   "TT426STR_ALM_ANALOG_DB_VERY LOW LEVEL VALUE (LL)" : Real = PLC TT426STR_ALM_ANALOG_DB."VERY LOW LEVEL VALUE (LL)" AT %DB2072.DBD22, 1 s
   "IDB_TIT 360_VERY HIGH LEVEL VALUE (HH)" : Real = PLC "IDB_TIT 360"."VERY HIGH LEVEL VALUE (HH)" AT %DB760.DBD34, 1 s
   "IDB_TIT 360_HIGH LEVEL VALUE (H)" : Real = PLC "IDB_TIT 360"."HIGH LEVEL VALUE (H)" AT %DB760.DBD30, 1 s
   "IDB_TIT 360_LOW LEVEL VALUE (L)" : Real = PLC "IDB_TIT 360"."LOW LEVEL VALUE (L)" AT %DB760.DBD26, 1 s
   "IDB_TIT 360_VERY LOW LEVEL VALUE (LL)" : Real = PLC "IDB_TIT 360"."VERY LOW LEVEL VALUE (LL)" AT %DB760.DBD22, 1 s
   "IDB_TIT 319_VERY HIGH LEVEL VALUE (HH)" : Real = PLC "IDB_TIT 319"."VERY HIGH LEVEL VALUE (HH)" AT %DB719.DBD34, 1 s
   "IDB_TIT 319_HIGH LEVEL VALUE (H)" : Real = PLC "IDB_TIT 319"."HIGH LEVEL VALUE (H)" AT %DB719.DBD30, 1 s
   "IDB_TIT 319_LOW LEVEL VALUE (L)" : Real = PLC "IDB_TIT 319"."LOW LEVEL VALUE (L)" AT %DB719.DBD26, 1 s
   "IDB_TIT 319_VERY LOW LEVEL VALUE (LL)" : Real = PLC "IDB_TIT 319"."VERY LOW LEVEL VALUE (LL)" AT %DB719.DBD22, 1 s
   "IDB_PIT 316_VERY HIGH LEVEL VALUE (HH)" : Real = PLC "IDB_PIT 316"."VERY HIGH LEVEL VALUE (HH)" AT %DB716.DBD34, 1 s
   "IDB_PIT 316_HIGH LEVEL VALUE (H)" : Real = PLC "IDB_PIT 316"."HIGH LEVEL VALUE (H)" AT %DB716.DBD30, 1 s
   "IDB_PIT 316_LOW LEVEL VALUE (L)" : Real = PLC "IDB_PIT 316"."LOW LEVEL VALUE (L)" AT %DB716.DBD26, 1 s
   "IDB_PIT 316_VERY LOW LEVEL VALUE (LL)" : Real = PLC "IDB_PIT 316"."VERY LOW LEVEL VALUE (LL)" AT %DB716.DBD22, 1 s
   "IDB_PIT 359_VERY HIGH LEVEL VALUE (HH)" : Real = PLC "IDB_PIT 359"."VERY HIGH LEVEL VALUE (HH)" AT %DB759.DBD34, 1 s
   "IDB_PIT 359_HIGH LEVEL VALUE (H)" : Real = PLC "IDB_PIT 359"."HIGH LEVEL VALUE (H)" AT %DB759.DBD30, 1 s
   "IDB_PIT 359_LOW LEVEL VALUE (L)" : Real = PLC "IDB_PIT 359"."LOW LEVEL VALUE (L)" AT %DB759.DBD26, 1 s
   "IDB_PIT 359_VERY LOW LEVEL VALUE (LL)" : Real = PLC "IDB_PIT 359"."VERY LOW LEVEL VALUE (LL)" AT %DB759.DBD22, 1 s
   "IDB_ATO2B_1_VERY HIGH LEVEL VALUE (HH)" : Real = PLC IDB_ATO2B_1."VERY HIGH LEVEL VALUE (HH)" AT %DB731.DBD34, 1 s
   "IDB_ATO2B_1_HIGH LEVEL VALUE (H)" : Real = PLC IDB_ATO2B_1."HIGH LEVEL VALUE (H)" AT %DB731.DBD30, 1 s
   "IDB_ATO2B_1_LOW LEVEL VALUE (L)" : Real = PLC IDB_ATO2B_1."LOW LEVEL VALUE (L)" AT %DB731.DBD26, 1 s
   "IDB_ATO2B_1_VERY LOW LEVEL VALUE (LL)" : Real = PLC IDB_ATO2B_1."VERY LOW LEVEL VALUE (LL)" AT %DB731.DBD22, 1 s
   "TT426_5S_ALM_ANALOG_DB_VERY HIGH LEVEL VALUE (HH)" : Real = PLC TT426_5S_ALM_ANALOG_DB."VERY HIGH LEVEL VALUE (HH)" AT %DB2082.DBD34, 1 s
   "TT426_5S_ALM_ANALOG_DB_HIGH LEVEL VALUE (H)" : Real = PLC TT426_5S_ALM_ANALOG_DB."HIGH LEVEL VALUE (H)" AT %DB2082.DBD30, 1 s
   "TT426_5S_ALM_ANALOG_DB_LOW LEVEL VALUE (L)" : Real = PLC TT426_5S_ALM_ANALOG_DB."LOW LEVEL VALUE (L)" AT %DB2082.DBD26, 1 s
   "TT426_5S_ALM_ANALOG_DB_VERY LOW LEVEL VALUE (LL)" : Real = PLC TT426_5S_ALM_ANALOG_DB."VERY LOW LEVEL VALUE (LL)" AT %DB2082.DBD22, 1 s
   "PIT424_RIO6_ALM_ANALOG_DB_VERY HIGH LEVEL VALUE (HH)" : Real = PLC PIT424_RIO6_ALM_ANALOG_DB."VERY HIGH LEVEL VALUE (HH)" AT %DB2223.DBD34, 1 s
   "PIT424_RIO6_ALM_ANALOG_DB_HIGH LEVEL VALUE (H)" : Real = PLC PIT424_RIO6_ALM_ANALOG_DB."HIGH LEVEL VALUE (H)" AT %DB2223.DBD30, 1 s
   "PIT424_RIO6_ALM_ANALOG_DB_LOW LEVEL VALUE (L)" : Real = PLC PIT424_RIO6_ALM_ANALOG_DB."LOW LEVEL VALUE (L)" AT %DB2223.DBD26, 1 s
   "PIT424_RIO6_ALM_ANALOG_DB_VERY LOW LEVEL VALUE (LL)" : Real = PLC PIT424_RIO6_ALM_ANALOG_DB."VERY LOW LEVEL VALUE (LL)" AT %DB2223.DBD22, 1 s
   "TT426_6P_ALM_ANALOG_DB_VERY HIGH LEVEL VALUE (HH)" : Real = PLC TT426_6P_ALM_ANALOG_DB."VERY HIGH LEVEL VALUE (HH)" AT %DB2083.DBD34, 1 s
   "TT426_6P_ALM_ANALOG_DB_HIGH LEVEL VALUE (H)" : Real = PLC TT426_6P_ALM_ANALOG_DB."HIGH LEVEL VALUE (H)" AT %DB2083.DBD30, 1 s
   "TT426_6P_ALM_ANALOG_DB_LOW LEVEL VALUE (L)" : Real = PLC TT426_6P_ALM_ANALOG_DB."LOW LEVEL VALUE (L)" AT %DB2083.DBD26, 1 s
   "TT426_6P_ALM_ANALOG_DB_VERY LOW LEVEL VALUE (LL)" : Real = PLC TT426_6P_ALM_ANALOG_DB."VERY LOW LEVEL VALUE (LL)" AT %DB2083.DBD22, 1 s
   "TT426_6S_ALM_ANALOG_DB_VERY HIGH LEVEL VALUE (HH)" : Real = PLC TT426_6S_ALM_ANALOG_DB."VERY HIGH LEVEL VALUE (HH)" AT %DB2085.DBD34, 1 s
   "TT426_6S_ALM_ANALOG_DB_HIGH LEVEL VALUE (H)" : Real = PLC TT426_6S_ALM_ANALOG_DB."HIGH LEVEL VALUE (H)" AT %DB2085.DBD30, 1 s
   "TT426_6S_ALM_ANALOG_DB_LOW LEVEL VALUE (L)" : Real = PLC TT426_6S_ALM_ANALOG_DB."LOW LEVEL VALUE (L)" AT %DB2085.DBD26, 1 s
   "TT426_6S_ALM_ANALOG_DB_VERY LOW LEVEL VALUE (LL)" : Real = PLC TT426_6S_ALM_ANALOG_DB."VERY LOW LEVEL VALUE (LL)" AT %DB2085.DBD22, 1 s
   "PIT424_RIO7_ALM_ANALOG_DB_VERY HIGH LEVEL VALUE (HH)" : Real = PLC PIT424_RIO7_ALM_ANALOG_DB."VERY HIGH LEVEL VALUE (HH)" AT %DB2224.DBD34, 1 s
   "PIT424_RIO7_ALM_ANALOG_DB_HIGH LEVEL VALUE (H)" : Real = PLC PIT424_RIO7_ALM_ANALOG_DB."HIGH LEVEL VALUE (H)" AT %DB2224.DBD30, 1 s
   "PIT424_RIO7_ALM_ANALOG_DB_LOW LEVEL VALUE (L)" : Real = PLC PIT424_RIO7_ALM_ANALOG_DB."LOW LEVEL VALUE (L)" AT %DB2224.DBD26, 1 s
   "PIT424_RIO7_ALM_ANALOG_DB_VERY LOW LEVEL VALUE (LL)" : Real = PLC PIT424_RIO7_ALM_ANALOG_DB."VERY LOW LEVEL VALUE (LL)" AT %DB2224.DBD22, 1 s
   "TT426_APT_ALM_ANALOG_DB_VERY HIGH LEVEL VALUE (HH)" : Real = PLC TT426_APT_ALM_ANALOG_DB."VERY HIGH LEVEL VALUE (HH)" AT %DB2087.DBD34, 1 s
   "TT426_APT_ALM_ANALOG_DB_HIGH LEVEL VALUE (H)" : Real = PLC TT426_APT_ALM_ANALOG_DB."HIGH LEVEL VALUE (H)" AT %DB2087.DBD30, 1 s
   "TT426_APT_ALM_ANALOG_DB_LOW LEVEL VALUE (L)" : Real = PLC TT426_APT_ALM_ANALOG_DB."LOW LEVEL VALUE (L)" AT %DB2087.DBD26, 1 s
   "TT426_APT_ALM_ANALOG_DB_VERY LOW LEVEL VALUE (LL)" : Real = PLC TT426_APT_ALM_ANALOG_DB."VERY LOW LEVEL VALUE (LL)" AT %DB2087.DBD22, 1 s
   "PIT424_RIO5_ALM_ANALOG_DB_VERY HIGH LEVEL VALUE (HH)" : Real = PLC PIT424_RIO5_ALM_ANALOG_DB."VERY HIGH LEVEL VALUE (HH)" AT %DB2222.DBD34, 1 s
   "PIT424_RIO5_ALM_ANALOG_DB_HIGH LEVEL VALUE (H)" : Real = PLC PIT424_RIO5_ALM_ANALOG_DB."HIGH LEVEL VALUE (H)" AT %DB2222.DBD30, 1 s
   "PIT424_RIO5_ALM_ANALOG_DB_LOW LEVEL VALUE (L)" : Real = PLC PIT424_RIO5_ALM_ANALOG_DB."LOW LEVEL VALUE (L)" AT %DB2222.DBD26, 1 s
   "PIT424_RIO5_ALM_ANALOG_DB_VERY LOW LEVEL VALUE (LL)" : Real = PLC PIT424_RIO5_ALM_ANALOG_DB."VERY LOW LEVEL VALUE (LL)" AT %DB2222.DBD22, 1 s
   "TT426_5P_ALM_ANALOG_DB_VERY HIGH LEVEL VALUE (HH)" : Real = PLC TT426_5P_ALM_ANALOG_DB."VERY HIGH LEVEL VALUE (HH)" AT %DB2081.DBD34, 1 s
   "TT426_5P_ALM_ANALOG_DB_HIGH LEVEL VALUE (H)" : Real = PLC TT426_5P_ALM_ANALOG_DB."HIGH LEVEL VALUE (H)" AT %DB2081.DBD30, 1 s
   "TT426_5P_ALM_ANALOG_DB_LOW LEVEL VALUE (L)" : Real = PLC TT426_5P_ALM_ANALOG_DB."LOW LEVEL VALUE (L)" AT %DB2081.DBD26, 1 s
   "TT426_5P_ALM_ANALOG_DB_VERY LOW LEVEL VALUE (LL)" : Real = PLC TT426_5P_ALM_ANALOG_DB."VERY LOW LEVEL VALUE (LL)" AT %DB2081.DBD22, 1 s
   "TT426_4S_ALM_ANALOG_DB_VERY HIGH LEVEL VALUE (HH)" : Real = PLC TT426_4S_ALM_ANALOG_DB."VERY HIGH LEVEL VALUE (HH)" AT %DB2080.DBD34, 1 s
   "TT426_4S_ALM_ANALOG_DB_HIGH LEVEL VALUE (H)" : Real = PLC TT426_4S_ALM_ANALOG_DB."HIGH LEVEL VALUE (H)" AT %DB2080.DBD30, 1 s
   "TT426_4S_ALM_ANALOG_DB_LOW LEVEL VALUE (L)" : Real = PLC TT426_4S_ALM_ANALOG_DB."LOW LEVEL VALUE (L)" AT %DB2080.DBD26, 1 s
   "TT426_4S_ALM_ANALOG_DB_VERY LOW LEVEL VALUE (LL)" : Real = PLC TT426_4S_ALM_ANALOG_DB."VERY LOW LEVEL VALUE (LL)" AT %DB2080.DBD22, 1 s
   "FIT419_ALM_ANALOG_DB_VERY HIGH LEVEL VALUE (HH)" : Real = PLC FIT419_ALM_ANALOG_DB."VERY HIGH LEVEL VALUE (HH)" AT %DB2067.DBD34, 1 s
   "FIT419_ALM_ANALOG_DB_HIGH LEVEL VALUE (H)" : Real = PLC FIT419_ALM_ANALOG_DB."HIGH LEVEL VALUE (H)" AT %DB2067.DBD30, 1 s
   "FIT419_ALM_ANALOG_DB_LOW LEVEL VALUE (L)" : Real = PLC FIT419_ALM_ANALOG_DB."LOW LEVEL VALUE (L)" AT %DB2067.DBD26, 1 s
   "FIT419_ALM_ANALOG_DB_VERY LOW LEVEL VALUE (LL)" : Real = PLC FIT419_ALM_ANALOG_DB."VERY LOW LEVEL VALUE (LL)" AT %DB2067.DBD22, 1 s
   "FIT417_2S_ALM_ANALOG_DB_VERY HIGH LEVEL VALUE (HH)" : Real = PLC FIT417_2S_ALM_ANALOG_DB."VERY HIGH LEVEL VALUE (HH)" AT %DB2066.DBD34, 1 s
   "FIT417_2S_ALM_ANALOG_DB_HIGH LEVEL VALUE (H)" : Real = PLC FIT417_2S_ALM_ANALOG_DB."HIGH LEVEL VALUE (H)" AT %DB2066.DBD30, 1 s
   "FIT417_2S_ALM_ANALOG_DB_LOW LEVEL VALUE (L)" : Real = PLC FIT417_2S_ALM_ANALOG_DB."LOW LEVEL VALUE (L)" AT %DB2066.DBD26, 1 s
   "FIT417_2S_ALM_ANALOG_DB_VERY LOW LEVEL VALUE (LL)" : Real = PLC FIT417_2S_ALM_ANALOG_DB."VERY LOW LEVEL VALUE (LL)" AT %DB2066.DBD22, 1 s
   "PIT424PORT_ALM_ANALOG_DB_HIGH LEVEL VALUE (H)" : Real = PLC PIT424PORT_ALM_ANALOG_DB."HIGH LEVEL VALUE (H)" AT %DB2070.DBD30, 1 s
   "PIT424PORT_ALM_ANALOG_DB_LOW LEVEL VALUE (L)" : Real = PLC PIT424PORT_ALM_ANALOG_DB."LOW LEVEL VALUE (L)" AT %DB2070.DBD26, 1 s
   "PIT424PORT_ALM_ANALOG_DB_VERY LOW LEVEL VALUE (LL)" : Real = PLC PIT424PORT_ALM_ANALOG_DB."VERY LOW LEVEL VALUE (LL)" AT %DB2070.DBD22, 1 s
   "FIT420PORT_ALM_ANALOG_DB_VERY HIGH LEVEL VALUE (HH)" : Real = PLC FIT420PORT_ALM_ANALOG_DB."VERY HIGH LEVEL VALUE (HH)" AT %DB2065.DBD34, 1 s
   "FIT420PORT_ALM_ANALOG_DB_HIGH LEVEL VALUE (H)" : Real = PLC FIT420PORT_ALM_ANALOG_DB."HIGH LEVEL VALUE (H)" AT %DB2065.DBD30, 1 s
   "FIT420PORT_ALM_ANALOG_DB_LOW LEVEL VALUE (L)" : Real = PLC FIT420PORT_ALM_ANALOG_DB."LOW LEVEL VALUE (L)" AT %DB2065.DBD26, 1 s
   "FIT420PORT_ALM_ANALOG_DB_VERY LOW LEVEL VALUE (LL)" : Real = PLC FIT420PORT_ALM_ANALOG_DB."VERY LOW LEVEL VALUE (LL)" AT %DB2065.DBD22, 1 s
   "FIT418_2P_ALM_ANALOG_DB_VERY HIGH LEVEL VALUE (HH)" : Real = PLC FIT418_2P_ALM_ANALOG_DB."VERY HIGH LEVEL VALUE (HH)" AT %DB2064.DBD34, 1 s
   "FIT418_2P_ALM_ANALOG_DB_HIGH LEVEL VALUE (H)" : Real = PLC FIT418_2P_ALM_ANALOG_DB."HIGH LEVEL VALUE (H)" AT %DB2064.DBD30, 1 s
   "FIT418_2P_ALM_ANALOG_DB_LOW LEVEL VALUE (L)" : Real = PLC FIT418_2P_ALM_ANALOG_DB."LOW LEVEL VALUE (L)" AT %DB2064.DBD26, 1 s
   "FIT418_2P_ALM_ANALOG_DB_VERY LOW LEVEL VALUE (LL)" : Real = PLC FIT418_2P_ALM_ANALOG_DB."VERY LOW LEVEL VALUE (LL)" AT %DB2064.DBD22, 1 s
   "PT415_RIO7_ALM_ANALOG_DB_VERY HIGH LEVEL VALUE (HH)" : Real = PLC PT415_RIO7_ALM_ANALOG_DB."VERY HIGH LEVEL VALUE (HH)" AT %DB2225.DBD34, 1 s
   "PT415_RIO7_ALM_ANALOG_DB_HIGH LEVEL VALUE (H)" : Real = PLC PT415_RIO7_ALM_ANALOG_DB."HIGH LEVEL VALUE (H)" AT %DB2225.DBD30, 1 s
   "PT415_RIO7_ALM_ANALOG_DB_LOW LEVEL VALUE (L)" : Real = PLC PT415_RIO7_ALM_ANALOG_DB."LOW LEVEL VALUE (L)" AT %DB2225.DBD26, 1 s
   "PT415_RIO7_ALM_ANALOG_DB_VERY LOW LEVEL VALUE (LL)" : Real = PLC PT415_RIO7_ALM_ANALOG_DB."VERY LOW LEVEL VALUE (LL)" AT %DB2225.DBD22, 1 s
   "PT415_RIO6_ALM_ANALOG_DB_VERY HIGH LEVEL VALUE (HH)" : Real = PLC PT415_RIO6_ALM_ANALOG_DB."VERY HIGH LEVEL VALUE (HH)" AT %DB2218.DBD34, 1 s
   "PT415_RIO6_ALM_ANALOG_DB_HIGH LEVEL VALUE (H)" : Real = PLC PT415_RIO6_ALM_ANALOG_DB."HIGH LEVEL VALUE (H)" AT %DB2218.DBD30, 1 s
   "PT415_RIO6_ALM_ANALOG_DB_LOW LEVEL VALUE (L)" : Real = PLC PT415_RIO6_ALM_ANALOG_DB."LOW LEVEL VALUE (L)" AT %DB2218.DBD26, 1 s
   "PT415_RIO6_ALM_ANALOG_DB_VERY LOW LEVEL VALUE (LL)" : Real = PLC PT415_RIO6_ALM_ANALOG_DB."VERY LOW LEVEL VALUE (LL)" AT %DB2218.DBD22, 1 s
   "PT415_RIO5_ALM_ANALOG_DB_VERY HIGH LEVEL VALUE (HH)" : Real = PLC PT415_RIO5_ALM_ANALOG_DB."VERY HIGH LEVEL VALUE (HH)" AT %DB2217.DBD34, 1 s
   "PT415_RIO5_ALM_ANALOG_DB_HIGH LEVEL VALUE (H)" : Real = PLC PT415_RIO5_ALM_ANALOG_DB."HIGH LEVEL VALUE (H)" AT %DB2217.DBD30, 1 s
   "PT415_RIO5_ALM_ANALOG_DB_LOW LEVEL VALUE (L)" : Real = PLC PT415_RIO5_ALM_ANALOG_DB."LOW LEVEL VALUE (L)" AT %DB2217.DBD26, 1 s
   "PT415_RIO5_ALM_ANALOG_DB_VERY LOW LEVEL VALUE (LL)" : Real = PLC PT415_RIO5_ALM_ANALOG_DB."VERY LOW LEVEL VALUE (LL)" AT %DB2217.DBD22, 1 s
   "PT415_RIO3_ALM_ANALOG_DB_VERY HIGH LEVEL VALUE (HH)" : Real = PLC PT415_RIO3_ALM_ANALOG_DB."VERY HIGH LEVEL VALUE (HH)" AT %DB2215.DBD34, 1 s
   "PT415_RIO3_ALM_ANALOG_DB_HIGH LEVEL VALUE (H)" : Real = PLC PT415_RIO3_ALM_ANALOG_DB."HIGH LEVEL VALUE (H)" AT %DB2215.DBD30, 1 s
   "PT415_RIO3_ALM_ANALOG_DB_LOW LEVEL VALUE (L)" : Real = PLC PT415_RIO3_ALM_ANALOG_DB."LOW LEVEL VALUE (L)" AT %DB2215.DBD26, 1 s
   "PT415_RIO3_ALM_ANALOG_DB_VERY LOW LEVEL VALUE (LL)" : Real = PLC PT415_RIO3_ALM_ANALOG_DB."VERY LOW LEVEL VALUE (LL)" AT %DB2215.DBD22, 1 s
   "PT415_FPT_ALM_ANALOG_DB_VERY HIGH LEVEL VALUE (HH)" : Real = PLC PT415_FPT_ALM_ANALOG_DB."VERY HIGH LEVEL VALUE (HH)" AT %DB2213.DBD34, 1 s
   "PT415_FPT_ALM_ANALOG_DB_HIGH LEVEL VALUE (H)" : Real = PLC PT415_FPT_ALM_ANALOG_DB."HIGH LEVEL VALUE (H)" AT %DB2213.DBD30, 1 s
   "PT415_FPT_ALM_ANALOG_DB_LOW LEVEL VALUE (L)" : Real = PLC PT415_FPT_ALM_ANALOG_DB."LOW LEVEL VALUE (L)" AT %DB2213.DBD26, 1 s
   "PT415_FPT_ALM_ANALOG_DB_VERY LOW LEVEL VALUE (LL)" : Real = PLC PT415_FPT_ALM_ANALOG_DB."VERY LOW LEVEL VALUE (LL)" AT %DB2213.DBD22, 1 s
   "Process Gas Compressor Running/Stopped" : Bool = PLC "Process Gas Compressor Running/Stopped" AT %I139.0, 1 s
   "504_Tank Grouping_DB2020_Valve Cycle_Enable" : Bool = PLC "504_Tank Grouping_DB2020"."Valve Cycle".Enable, 1 s
   "504_Tank Grouping_DB2020_Valve Cycle_Period" : Time = PLC "504_Tank Grouping_DB2020"."Valve Cycle".Period, 1 s
   "504_Tank Grouping_DB2020_Valve Cycle_Length" : Time = PLC "504_Tank Grouping_DB2020"."Valve Cycle".Length, 1 s
   "504_Tank Grouping_DB2020_Cycle Period_ET" : Time = PLC "504_Tank Grouping_DB2020"."Cycle Period".ET, 1 s
   "504_Tank Grouping_DB2020_Cycle Length_ET" : Time = PLC "504_Tank Grouping_DB2020"."Cycle Length".ET, 1 s
   "Sequence Times_DB_Jurney Time FB_Hours Left" : Int = PLC "Sequence Times_DB"."Jurney Time FB"."Hours Left", 1 s
   "Sequence Times_DB_Jurney Time FB_Days Left" : Int = PLC "Sequence Times_DB"."Jurney Time FB"."Days Left", 1 s
   "Sequence Times_DB_Pre-Dwell Timer_Minutes Left" : DInt = PLC "Sequence Times_DB"."Pre-Dwell Timer"."Minutes Left", 1 s
   "Sequence Times_DB_Pre-Dwell Timer_Hours Left" : DInt = PLC "Sequence Times_DB"."Pre-Dwell Timer"."Hours Left", 1 s
   "Sequence Times_DB_Pre-Dwell Timer_Days Left" : DInt = PLC "Sequence Times_DB"."Pre-Dwell Timer"."Days Left", 1 s
   "Sequence Times_DB_Jurney Time" : Real = PLC "Sequence Times_DB"."Jurney Time", 1 s
   "Sequence Times_DB_Treatment Timer_Days" : DInt = PLC "Sequence Times_DB"."Treatment Timer".Days, 1 s
   "Sequence Times_DB_Treatment Timer_Hours" : DInt = PLC "Sequence Times_DB"."Treatment Timer".Hours, 1 s
   "Sequence Times_DB_Treatment Timer_Minutes" : DInt = PLC "Sequence Times_DB"."Treatment Timer".Minutes, 1 s
   "Sequence Times_DB_Treatment Timer_Days Left" : DInt = PLC "84_Setpoints".PIT113_Low, 1 s
   "Sequence Times_DB_Treatment Timer_Hours Left" : DInt = PLC "Sequence Times_DB"."Treatment Timer"."Hours Left", 1 s
   "Sequence Times_DB_Treatment Timer_Minutes Left" : DInt = PLC "Sequence Times_DB"."Treatment Timer"."Minutes Left", 1 s
   "Sequence Times_DB_Pre-Dwell Timer_PT_HOURS" : Real = PLC "Sequence Times_DB"."Pre-Dwell Timer".PT_HOURS, 1 s
   "Sequence Times_DB_De-Ox Timer_PT_HOURS" : Real = PLC "Sequence Times_DB"."De-Ox Timer".PT_HOURS, 1 s
   "Sequence Times_DB_De-Ox Timer_Days Left" : DInt = PLC "Sequence Times_DB"."De-Ox Timer"."Days Left", 1 s
   "Sequence Times_DB_De-Ox Timer_Hours Left" : DInt = PLC "Sequence Times_DB"."De-Ox Timer"."Hours Left", 1 s
   "Sequence Times_DB_De-Ox Timer_Minutes Left" : DInt = PLC "Sequence Times_DB"."De-Ox Timer"."Minutes Left", 1 s
   "504_Tank Grouping_DB2020_O2 De-Ox Setpoint" : Real = PLC "504_Tank Grouping_DB2020"."O2 De-Ox Setpoint", 1 s
   "Sequence Times_DB_Dwell Timer_PT_HOURS" : Real = PLC "Sequence Times_DB"."Dwell Timer".PT_HOURS, 1 s
   "Sequence Times_DB_Dwell Timer_Days Left" : DInt = PLC "Sequence Times_DB"."Dwell Timer"."Days Left", 1 s
   "Sequence Times_DB_Dwell Timer_Hours Left" : DInt = PLC "Sequence Times_DB"."Dwell Timer"."Hours Left", 1 s
   "Sequence Times_DB_Dwell Timer_Minutes Left" : DInt = PLC "Sequence Times_DB"."Dwell Timer"."Minutes Left", 1 s
   "Sequence Times_DB_Re-Ox Timer_PT_HOURS" : Real = PLC "Sequence Times_DB"."Re-Ox Timer".PT_HOURS, 1 s
   "Sequence Times_DB_Re-Ox Timer_Days Left" : DInt = PLC "Sequence Times_DB"."Re-Ox Timer"."Days Left", 1 s
   "Sequence Times_DB_Re-Ox Timer_Hours Left" : DInt = PLC "Sequence Times_DB"."Re-Ox Timer"."Hours Left", 1 s
   "Sequence Times_DB_Re-Ox Timer_Minutes Left" : DInt = PLC "Sequence Times_DB"."Re-Ox Timer"."Minutes Left", 1 s
   "Sequence Times_DB_Post-Dwell Timer_PT_HOURS" : Real = PLC "Sequence Times_DB"."Post-Dwell Timer".PT_HOURS, 1 s
   "Sequence Times_DB_Post-Dwell Timer_Days Left" : DInt = PLC "Sequence Times_DB"."Post-Dwell Timer"."Days Left", 1 s
   "Sequence Times_DB_Post-Dwell Timer_Hours Left" : DInt = PLC "Sequence Times_DB"."Post-Dwell Timer"."Hours Left", 1 s
   "Sequence Times_DB_Post-Dwell Timer_Minutes Left" : DInt = PLC "Sequence Times_DB"."Post-Dwell Timer"."Minutes Left", 1 s
   "Sequence Times_DB_Pre-Dwell Time" : Real = PLC "Sequence Times_DB"."Pre-Dwell Time", 1 s
   "Sequence Times_DB_De-Ox Time" : Real = PLC "Sequence Times_DB"."De-Ox Time", 1 s
   "Sequence Times_DB_De-Ox SP Time" : Real = PLC "Sequence Times_DB"."De-Ox SP Time", 1 s
   "Sequence Times_DB_Dwell Time" : Real = PLC "Sequence Times_DB"."Dwell Time", 1 s
   "Sequence Times_DB_Re-Ox Time" : Real = PLC "Sequence Times_DB"."Re-Ox Time", 1 s
   "Sequence Times_DB_Post-Dwell Time" : Real = PLC "Sequence Times_DB"."Post-Dwell Time", 1 s
   "2068_Sys_Status_Data_Not BWT mode Warning" : Bool = PLC "2068_Sys_Status_Data"."Not BWT mode Warning" AT %DB1.DBX0.0, 1 s
      on ChangeValue: "BWT_Warning"()
   "2086_Times_CV422_FPT_MAX_TRVL_TIME" : Time = PLC "2086_Times".CV422_FPT_MAX_TRVL_TIME, 1 s
   "2086_Times_CV422_1P_MAX_TRVL_TIME" : Time = PLC "2086_Times".CV422_1P_MAX_TRVL_TIME, 1 s
   "2086_Times_CV421_1S_MAX_TRVL_TIME" : Time = PLC "2086_Times".CV421_1S_MAX_TRVL_TIME, 1 s
   "2086_Times_CV422_2P_MAX_TRVL_TIME" : Time = PLC "2086_Times".CV422_2P_MAX_TRVL_TIME, 1 s
   "2086_Times_CV421_2S_MAX_TRVL_TIME" : Time = PLC "2086_Times".CV421_2S_MAX_TRVL_TIME, 1 s
   "2086_Times_CV422_3P_MAX_TRVL_TIME" : Time = PLC "2086_Times".CV422_3P_MAX_TRVL_TIME, 1 s
   "2086_Times_CV421_3S_MAX_TRVL_TIME" : Time = PLC "2086_Times".CV421_3S_MAX_TRVL_TIME, 1 s
   "2086_Times_CV422_4P_MAX_TRVL_TIME" : Time = PLC "2086_Times".CV422_4P_MAX_TRVL_TIME, 1 s
   "2086_Times_CV421_4S_MAX_TRVL_TIME" : Time = PLC "2086_Times".CV421_4S_MAX_TRVL_TIME, 1 s
   "2086_Times_CV422_5P_MAX_TRVL_TIME" : Time = PLC "2086_Times".CV422_5P_MAX_TRVL_TIME, 1 s
   "2086_Times_CV421_5S_MAX_TRVL_TIME" : Time = PLC "2086_Times".CV421_5S_MAX_TRVL_TIME, 1 s
   "2086_Times_CV422_6P_MAX_TRVL_TIME" : Time = PLC "2086_Times".CV422_6P_MAX_TRVL_TIME, 1 s
   "2086_Times_CV421_6S_MAX_TRVL_TIME" : Time = PLC "2086_Times".CV421_6S_MAX_TRVL_TIME, 1 s
   "2086_Times_CV422_APT_MAX_TRVL_TIME" : Time = PLC "2086_Times".CV422_APT_MAX_TRVL_TIME, 1 s
   "Sequence Times_DB_Treatment Timer_Enable" : Bool = PLC "Sequence Times_DB"."Treatment Timer".Enable, 1 s
   "504_Tank Grouping_DB2020_Sequence Time m Offset_Int" : Real = PLC "504_Tank Grouping_DB2020"."Sequence Time m Offset_real", 1 s
   "504_Tank Grouping_DB2020_Boost" : Bool = PLC "504_Tank Grouping_DB2020".Boost, 1 s
   "503_WARNING CHCK_DB_2063_Alarm Word 12" : Word = PLC "503_WARNING CHCK_DB_2063"."Alarm Word 12", 1 s
   "503_WARNING CHCK_DB_2063_Alarm Word 13" : Word = PLC "503_WARNING CHCK_DB_2063"."Alarm Word 13", 1 s
   "503_WARNING CHCK_DB_2063_Alarm Word 14" : Word = PLC "503_WARNING CHCK_DB_2063"."Alarm Word 14", 1 s
   "503_WARNING CHCK_DB_2063_Alarm Word 15" : Word = PLC "503_WARNING CHCK_DB_2063"."Alarm Word 15", 1 s
   "503_WARNING CHCK_DB_2063_Alarm Word 16" : Word = PLC "84_Setpoints"."E-400 PT002 Tolerance", 1 s
   "2062_Warning_Data_BTCS_WARNING_WORD_12" : Word = PLC "2062_Warning_Data".BTCS_WARNING_WORD_12 AT %DB2062.DBW362, 1 s
   "2062_Warning_Data_BTCS_WARNING_WORD_13" : Word = PLC "2062_Warning_Data".BTCS_WARNING_WORD_13 AT %DB2062.DBW364, 1 s
   "2062_Warning_Data_BTCS_WARNING_WORD_14" : Word = PLC "2062_Warning_Data".BTCS_WARNING_WORD_14 AT %DB2062.DBW366, 1 s
   "2062_Warning_Data_BTCS_WARNING_WORD_15" : Word = PLC "2062_Warning_Data".BTCS_WARNING_WORD_15 AT %DB2062.DBW368, 1 s
   "2062_Warning_Data_BTCS_WARNING_WORD_16" : Word = PLC "2062_Warning_Data".BTCS_WARNING_WORD_16 AT %DB2062.DBW370, 1 s
   "Sequence Times_DB_Warn to IGG Start" : Bool = PLC "Sequence Times_DB"."Warn to IGG Start" AT %DB1.DBW0, 1 s
      on ChangeValue: "TimeRemainingToTreatment"()
   "Sequence Times_DB_Pre-Dwell Timer_PT_DAYS" : Real = PLC "Sequence Times_DB"."Pre-Dwell Timer".PT_DAYS, 1 s
   "Sequence Times_DB_Pre-Dwell Timer_PT_MINUTES" : Real = PLC "Sequence Times_DB"."Pre-Dwell Timer".PT_MINUTES, 1 s
   "Sequence Times_DB_Jurney Time FB_PT_DAYS" : Real = PLC "Sequence Times_DB"."Jurney Time FB".PT_DAYS, 1 s
   "Sequence Times_DB_Jurney Timer_PT_DAYS" : Real = PLC "Sequence Times_DB"."Jurney Timer".PT_DAYS, 1 s
   "Sequence Times_DB_Jurney Timer_PT_HOURS" : Real = PLC "Sequence Times_DB"."Jurney Timer".PT_HOURS, 1 s
   "Sequence Times_DB_Jurney Timer_PT_MINUTES" : Real = PLC "Sequence Times_DB"."Jurney Timer".PT_MINUTES, 1 s
   "2068_Sys_Status_Data_Not BWT mode Warning(1)" : Bool = PLC "2068_Sys_Status_Data"."Not BWT mode Warning" AT %DB1.DBD0, 1 s
   "Sequence Times_DB_Continue" : Bool = PLC "Sequence Times_DB".Continue, 1 s
   "Recipe Tag" : Int AT %DB1.DBX0.0
   "Record Data Tag" : Int AT %DB1.DBX0.0
   "Data_From_WBT_Level_APT" : Real = PLC Data_From_WBT.Level_APT, 1 s
   "Data_From_WBT_Level_WBT_6P" : Real = PLC Data_From_WBT.Level_WBT_6P, 1 s
   "Data_From_WBT_Level_WBT_5P" : Real = PLC Data_From_WBT.Level_WBT_5P, 1 s
   "Data_From_WBT_Level_WBT_4P" : Real = PLC Data_From_WBT.Level_WBT_4P, 1 s
   "Data_From_WBT_Level_WBT_3P" : Real = PLC Data_From_WBT.Level_WBT_3P, 1 s
   "Data_From_WBT_Level_WBT_2P" : Real = PLC Data_From_WBT.Level_WBT_2P, 1 s
   "Data_From_WBT_Level_WBT_1P" : Real = PLC Data_From_WBT.Level_WBT_1P, 1 s
   "Data_From_WBT_Level_FPT" : Real = PLC Data_From_WBT.Level_FPT, 1 s
   "Data_From_WBT_Level_WBT_1S" : Real = PLC Data_From_WBT.Level_WBT_1S, 1 s
   "Data_From_WBT_Level_WBT_2S" : Real = PLC Data_From_WBT.Level_WBT_2S, 1 s
   "Data_From_WBT_Level_WBT_3S" : Real = PLC Data_From_WBT.Level_WBT_3S, 1 s
   "Data_From_WBT_Level_WBT_4S" : Real = PLC Data_From_WBT.Level_WBT_4S, 1 s
   "Data_From_WBT_Level_WBT_5S" : Real = PLC Data_From_WBT.Level_WBT_5S, 1 s
   "Data_From_WBT_Level_WBT_6S" : Real = PLC Data_From_WBT.Level_WBT_6S, 1 s
   "IN_Level_APT" : Int = PLC IN_Level_APT AT %IW1026, 1 s
   "Data_From_WBT_Level_APT m" : Real = PLC Data_From_WBT."Level_APT m", 1 s
   "Data_From_WBT_Level_WBT_6S m" : Real = PLC Data_From_WBT."Level_WBT_6S m", 1 s
   "Data_From_WBT_Level_WBT_5S m" : Real = PLC Data_From_WBT."Level_WBT_5S m", 1 s
   "Data_From_WBT_Level_WBT_4S m" : Real = PLC Data_From_WBT."Level_WBT_4S m", 1 s
   "Data_From_WBT_Level_WBT_3S m" : Real = PLC Data_From_WBT."Level_WBT_3S m", 1 s
   "Data_From_WBT_Level_WBT_2S m" : Real = PLC Data_From_WBT."Level_WBT_2S m", 1 s
   "Data_From_WBT_Level_WBT_1S m" : Real = PLC Data_From_WBT."Level_WBT_1S m", 1 s
   "Data_From_WBT_Level_FPT m" : Real = PLC Data_From_WBT."Level_FPT m", 1 s
   "Data_From_WBT_Level_WBT_1P m" : Real = PLC Data_From_WBT."Level_WBT_1P m", 1 s
   "Data_From_WBT_Level_WBT_2P m" : Real = PLC Data_From_WBT."Level_WBT_2P m", 1 s
   "Data_From_WBT_Level_WBT_3P m" : Real = PLC Data_From_WBT."Level_WBT_3P m", 1 s
   "Data_From_WBT_Level_WBT_4P m" : Real = PLC Data_From_WBT."Level_WBT_4P m", 1 s
   "Data_From_WBT_Level_WBT_5P m" : Real = PLC Data_From_WBT."Level_WBT_5P m", 1 s
   "Data_From_WBT_Level_WBT_6P m" : Real = PLC Data_From_WBT."Level_WBT_6P m", 1 s
   "E-400 Animation_DB_Animation" : Int = PLC "E-400 Animation_DB".Animation, 1 s
   "CSW_Animation_DB_Animation" : Int = PLC CSW_Animation_DB.Animation, 1 s
   "504_Tank Grouping_DB2020_Time Left Tank_Time Left m Tank 1" : DInt = PLC "504_Tank Grouping_DB2020"."Time Left Tank"."Time Left m Tank 1", 1 s
   "504_Tank Grouping_DB2020_Time Left Tank_Time Left h Tank 1" : DInt = PLC "504_Tank Grouping_DB2020"."Time Left Tank"."Time Left h Tank 1", 1 s
   "504_Tank Grouping_DB2020_Time Left Tank_Time Left d Tank 1" : DInt = PLC "504_Tank Grouping_DB2020"."Time Left Tank"."Time Left d Tank 1", 1 s
   "504_Tank Grouping_DB2020_Time Left Tank_Time Left m Tank 2" : DInt = PLC "504_Tank Grouping_DB2020"."Time Left Tank"."Time Left m Tank 2", 1 s
   "504_Tank Grouping_DB2020_Time Left Tank_Time Left h Tank 14" : DInt = PLC "504_Tank Grouping_DB2020"."Time Left Tank"."Time Left h Tank 14", 1 s
   "504_Tank Grouping_DB2020_Time Left Tank_Time Left d Tank 14" : DInt = PLC "504_Tank Grouping_DB2020"."Time Left Tank"."Time Left d Tank 14", 1 s
   "504_Tank Grouping_DB2020_Time Left Tank_Time Left m Tank 14" : DInt = PLC "504_Tank Grouping_DB2020"."Time Left Tank"."Time Left m Tank 14", 1 s
   "504_Tank Grouping_DB2020_Time Left Tank_Time Left h Tank 2" : DInt = PLC "504_Tank Grouping_DB2020"."Time Left Tank"."Time Left h Tank 2", 1 s
   "504_Tank Grouping_DB2020_Time Left Tank_Time Left d Tank 2" : DInt = PLC "504_Tank Grouping_DB2020"."Time Left Tank"."Time Left d Tank 2", 1 s
   "504_Tank Grouping_DB2020_Time Left Tank_Time Left m Tank 3" : DInt = PLC "504_Tank Grouping_DB2020"."Time Left Tank"."Time Left m Tank 3", 1 s
   "504_Tank Grouping_DB2020_Time Left Tank_Time Left h Tank 3" : DInt = PLC "504_Tank Grouping_DB2020"."Time Left Tank"."Time Left h Tank 3", 1 s
   "504_Tank Grouping_DB2020_Time Left Tank_Time Left d Tank 3" : DInt = PLC "504_Tank Grouping_DB2020"."Time Left Tank"."Time Left d Tank 3", 1 s
   "504_Tank Grouping_DB2020_Time Left Tank_Time Left m Tank 4" : DInt = PLC "504_Tank Grouping_DB2020"."Time Left Tank"."Time Left m Tank 4", 1 s
   "504_Tank Grouping_DB2020_Time Left Tank_Time Left h Tank 4" : DInt = PLC "LT422 4P  TANK LEVEL ALARM"."VERY LOW LEVEL VALUE (LL)", 1 s
   "504_Tank Grouping_DB2020_Time Left Tank_Time Left d Tank 4" : DInt = PLC "504_Tank Grouping_DB2020"."Time Left Tank"."Time Left d Tank 4", 1 s
   "504_Tank Grouping_DB2020_Time Left Tank_Time Left m Tank 5" : DInt = PLC "504_Tank Grouping_DB2020"."Time Left Tank"."Time Left m Tank 5", 1 s
   "504_Tank Grouping_DB2020_Time Left Tank_Time Left h Tank 5" : DInt = PLC "504_Tank Grouping_DB2020"."Time Left Tank"."Time Left h Tank 5", 1 s
   "504_Tank Grouping_DB2020_Time Left Tank_Time Left d Tank 5" : DInt = PLC "504_Tank Grouping_DB2020"."Time Left Tank"."Time Left d Tank 5", 1 s
   "504_Tank Grouping_DB2020_Time Left Tank_Time Left m Tank 6" : DInt = PLC "504_Tank Grouping_DB2020"."Time Left Tank"."Time Left m Tank 6", 1 s
   "504_Tank Grouping_DB2020_Time Left Tank_Time Left h Tank 6" : DInt = PLC "504_Tank Grouping_DB2020"."Time Left Tank"."Time Left h Tank 6", 1 s
   "504_Tank Grouping_DB2020_Time Left Tank_Time Left d Tank 6" : DInt = PLC "504_Tank Grouping_DB2020"."Time Left Tank"."Time Left d Tank 6", 1 s
   "504_Tank Grouping_DB2020_Time Left Tank_Time Left m Tank 7" : DInt = PLC "504_Tank Grouping_DB2020"."Time Left Tank"."Time Left m Tank 7", 1 s
   "504_Tank Grouping_DB2020_Time Left Tank_Time Left h Tank 7" : DInt = PLC "504_Tank Grouping_DB2020"."Time Left Tank"."Time Left h Tank 7", 1 s
   "504_Tank Grouping_DB2020_Time Left Tank_Time Left d Tank 7" : DInt = PLC "504_Tank Grouping_DB2020"."Time Left Tank"."Time Left d Tank 7", 1 s
   "504_Tank Grouping_DB2020_Time Left Tank_Time Left m Tank 8" : DInt = PLC "504_Tank Grouping_DB2020"."Time Left Tank"."Time Left m Tank 8", 1 s
   "504_Tank Grouping_DB2020_Time Left Tank_Time Left h Tank 8" : DInt = PLC "504_Tank Grouping_DB2020"."Time Left Tank"."Time Left h Tank 8", 1 s
   "504_Tank Grouping_DB2020_Time Left Tank_Time Left d Tank 8" : DInt = PLC "504_Tank Grouping_DB2020"."Time Left Tank"."Time Left d Tank 8", 1 s
   "504_Tank Grouping_DB2020_Time Left Tank_Time Left m Tank 9" : DInt = PLC "504_Tank Grouping_DB2020"."Time Left Tank"."Time Left m Tank 9", 1 s
   "504_Tank Grouping_DB2020_Time Left Tank_Time Left h Tank 9" : DInt = PLC "504_Tank Grouping_DB2020"."Time Left Tank"."Time Left h Tank 9", 1 s
   "504_Tank Grouping_DB2020_Time Left Tank_Time Left d Tank 9" : DInt = PLC "504_Tank Grouping_DB2020"."Time Left Tank"."Time Left d Tank 9", 1 s
   "504_Tank Grouping_DB2020_Time Left Tank_Time Left m Tank 10" : DInt = PLC "504_Tank Grouping_DB2020"."Time Left Tank"."Time Left m Tank 10", 1 s
   "504_Tank Grouping_DB2020_Time Left Tank_Time Left h Tank 10" : DInt = PLC "504_Tank Grouping_DB2020"."Time Left Tank"."Time Left h Tank 10", 1 s
   "504_Tank Grouping_DB2020_Time Left Tank_Time Left d Tank 10" : DInt = PLC "504_Tank Grouping_DB2020"."Time Left Tank"."Time Left d Tank 10", 1 s
   "504_Tank Grouping_DB2020_Time Left Tank_Time Left m Tank 11" : DInt = PLC "504_Tank Grouping_DB2020"."Time Left Tank"."Time Left m Tank 11", 1 s
   "504_Tank Grouping_DB2020_Time Left Tank_Time Left h Tank 11" : DInt = PLC "2084_Setpoints"."TX427 Star DO High", 1 s
   "504_Tank Grouping_DB2020_Time Left Tank_Time Left d Tank 11" : DInt = PLC "504_Tank Grouping_DB2020"."Time Left Tank"."Time Left d Tank 11", 1 s
   "504_Tank Grouping_DB2020_Time Left Tank_Time Left m Tank 12" : DInt = PLC "504_Tank Grouping_DB2020"."Time Left Tank"."Time Left m Tank 12", 1 s
   "504_Tank Grouping_DB2020_Time Left Tank_Time Left h Tank 12" : DInt = PLC "504_Tank Grouping_DB2020"."Time Left Tank"."Time Left h Tank 12", 1 s
   "504_Tank Grouping_DB2020_Time Left Tank_Time Left d Tank 12" : DInt = PLC "504_Tank Grouping_DB2020"."Time Left Tank"."Time Left d Tank 12", 1 s
   "504_Tank Grouping_DB2020_Time Left Tank_Time Left m Tank 13" : DInt = PLC "504_Tank Grouping_DB2020"."Time Left Tank"."Time Left m Tank 13", 1 s
   "504_Tank Grouping_DB2020_Time Left Tank_Time Left h Tank 13" : DInt = PLC "504_Tank Grouping_DB2020"."Time Left Tank"."Time Left h Tank 13", 1 s
   "504_Tank Grouping_DB2020_Time Left Tank_Time Left d Tank 13" : DInt = PLC "504_Tank Grouping_DB2020"."Time Left Tank"."Time Left d Tank 13", 1 s
   "PGC Flush_DB_PGC Stop Delay" : Time = PLC "PGC Flush_DB"."PGC Stop Delay", 1 s
   "PGC Flush_DB_CAB after Start Delay" : Time = PLC "PGC Flush_DB"."CAB after Start Delay", 1 s
   "PGC Flush_DB_CAB RPM Cmnd" : Real = PLC "PGC Flush_DB"."CAB RPM Cmd", 1 s
   "PGC Flush_DB_Override" : Bool = PLC "PGC Flush_DB".Override, 1 s
   "PGC Flush_DB_Running" : Bool = PLC "PGC Flush_DB".Running, 1 s
   "PGC Flush_DB_Activate" : Bool = PLC "PGC Flush_DB".Activate, 1 s
   "PGC Flush_DB_Done" : Bool = PLC "PGC Flush_DB".Done, 1 s
   "PGC Flush_DB_CV405 Open" : Bool = PLC "PGC Flush_DB"."CV405 Open", 1 s
   "PGC Flush_DB_CV401 Open" : Bool = PLC "PGC Flush_DB"."CV401 Open", 1 s
   "PGC Flush_DB_CV431 Open" : Bool = PLC "PGC Flush_DB"."CV431 Open", 1 s
   "PGC Flush_DB_CAB Start" : Bool = PLC "19_AUTO_CMNDS_Data".PIT353_CMND_LowLow, 1 s
   "PGC Flush_DB_CV403 Modulate" : Bool = PLC "PGC Flush_DB"."CV403 Modulate", 1 s
   "PGC Flush_DB_Stop PGC" : Bool = PLC "PGC Flush_DB"."Stop PGC", 1 s
   "PGC Flush_DB_PGC Purge Duration" : Time = PLC "PGC Flush_DB"."PGC Purge Duration", 1 s
   "PGC Flush_DB_CV403 Open" : Bool = PLC "PGC Flush_DB"."CV403 Open", 1 s
   "PGC Flush_DB_Flip Flop_Override_Output" : Bool = PLC "PGC Flush_DB"."Flip Flop_Override".Output, 1 s
   "19_AUTO_CMNDS_Data_Purge Rqst Simulate" : Bool = PLC "19_AUTO_CMNDS_Data"."Purge Rqst Simulate", 1 s
   "1405_PID_CV405_ManualEnable" : Bool = PLC "1405_PID_CV405".ManualEnable, 1 s
   "PGC Flush_DB_CV401 Opened" : Bool = PLC "PGC Flush_DB"."CV401 Opened", 1 s
   "PGC Flush_DB_CV431 Opened" : Bool = PLC "PGC Flush_DB"."CV431 Opened", 1 s
   "PGC Flush_DB_CV441 Closed" : Bool = PLC "PGC Flush_DB"."CV441 Closed", 1 s
   "PGC Flush_DB_CAB Started" : Bool = PLC "PGC Flush_DB"."CAB Started", 1 s
   "1403_PID_300CV403_ModeActivate" : Bool = PLC "1403_PID_300CV403".ModeActivate, 1 s
   "PGC Flush_DB_PGC Stoped" : Bool = PLC "PGC Flush_DB"."PGC Stoped", 1 s
   "1403_PID_300CV403_ManualEnable" : Bool = PLC "1403_PID_300CV403".ManualEnable, 1 s
   "20_TANKS_IP_DATA_RIO_01_SECOND_TANK_DECK_IG_PRESS" : Real = PLC "20_TANKS_IP_DATA".RIO_01.SECOND_TANK.DECK_IG_PRESS, 1 s
   "20_TANKS_IP_DATA_RIO_01_SECOND_TANK_O2_MONITOR" : Real = PLC "20_TANKS_IP_DATA".RIO_01.SECOND_TANK.O2_MONITOR, 1 s
   "20_TANKS_IP_DATA_RIO_03_SECOND_TANK_DECK_IG_PRESS" : Real = PLC "20_TANKS_IP_DATA".RIO_03.SECOND_TANK.DECK_IG_PRESS, 1 s
   "20_TANKS_IP_DATA_RIO_04_SECOND_TANK_DECK_IG_PRESS" : Real = PLC "20_TANKS_IP_DATA".RIO_04.SECOND_TANK.DECK_IG_PRESS, 1 s
   "20_TANKS_IP_DATA_RIO_05_SECOND_TANK_DECK_IG_PRESS" : Real = PLC "20_TANKS_IP_DATA".RIO_05.SECOND_TANK.DECK_IG_PRESS, 1 s
   "20_TANKS_IP_DATA_RIO_06_SECOND_TANK_DECK_IG_PRESS" : Real = PLC "20_TANKS_IP_DATA".RIO_06.SECOND_TANK.DECK_IG_PRESS, 1 s
   "20_TANKS_IP_DATA_RIO_06_SECOND_TANK_O2_MONITOR" : Real = PLC "20_TANKS_IP_DATA".RIO_06.SECOND_TANK.O2_MONITOR, 1 s
   "LOG IGG" : Bool = PLC "68_Sys_Status_Data"."LOG IGG" AT %DB1.DBW0, 1 s
      on ChangeValue: function_fd9437ed(0, "IGG_BC_FD001_Flame Detector"); function_fd9437ed(0, "GCU_FW_TIT408_Fresh water cooling"); function_fd9437ed(0, "IGG_Fuel_TIT202_Fuel Oil"); function_fd9437ed(0, "IGG_IG_TIT401_IG vent"); function_fd9437ed(0, "IGG_SW_TIT319_Cooling water (main line)"); function_fd9437ed(0, "IGG_SW_TIT360_Cooling water to drain line"); function_fd9437ed(0, "IGG_SW_TIT315_CW Temp to IGG Jacket"); function_fd9437ed(0, "IGG_CAB_PIT102_Comb Air"); function_fd9437ed(0, "IGG_Fuel_PIT204_Fuel Oil"); function_fd9437ed(0, "IGG_IA_PIT113_Atom Air to MBurner"); function_fd9437ed(0, "IGG_Fuel_PIT205_Fuel to MBurner"); function_fd9437ed(0, "IGG_IG_PIT402_IG vent"); function_fd9437ed(0, "IGG_SW_PIT359_Cooling water (main line)"); function_fd9437ed(0, "IGG_IA_PIT112_Inst Air"); function_fd9437ed(0, "IGG_SW_PIT316_Cooling water to IGG Jacket"); function_fd9437ed(0, "IGG_IG_TX-431_Atm Oxygen 1")